
screen "Air System" 1280x800, template "Template"
   Button "Button_16" at 609,168 size 64x25; TextOn 'Alarm'; TextOff 'Text'
   Button "Button_2" at 602,168 size 71x25; TextOn 'Alarm'; TextOff 'Shutdown'
      Visibility <- "10 DI_DATA_E131_SHTDN"
   Button "HmiScreenItemData_1" at 1,1 size 150x43; TextOn 'Back'; TextOff 'Main Index'
      on Release: ActivateScreen("02 Main Index", 0)
   Button "Button_15" at 464,168 size 57x25; TextOn 'Enabled'; TextOff 'Disabled'
   TextField "Text field_14" at 307,171 size 158x18; Text 'I & A Air Compressor'
   TextField "Text field_15" at 464,146 size 60x18; Text 'Enabled'
   TextField "Text field_16" at 530,146 size 64x18; Text 'Running'
   TextField "Text field_18" at 601,145 size 78x18; Text 'Shutdown'
   Button "Button_1" at 530,168 size 57x25; TextOn 'Enabled'; TextOff 'Stopped'
   TextField "Text field_1" at 282,55 size 561x26; Text 'Instrument & Atomising Air Compressor Control (E-131)'
   TextField "Text field_32" at 464,168 size 57x25; Text 'Enabled'
      Visibility <- "14_DQ_Data_E131ControlOut"
   TextField "Text field_2" at 530,168 size 57x25; Text 'Running'
      Visibility <- "10 DI_DATA_E131_OK"
   GraphicIOField "Graphic I/O field_2" at 703,308 size 196x199; PictureList "IA Compressor_2"
      ProcessValue <- "82_To_HMI_CA Blower Animation"
   Gauge "Gauge_1" at 791,570 size 184x184; CaptionText 'Open'; UnitText '%'
      ProcessValue <- "12_AI_Data_CV403_SCALED"
   TextField "Text field_20" at 374,532 size 529x26; Text 'Combustion Air/Inert Gas Pressure Control (CV-403)'
   IOField "I/O field_16" at 516,441 size 74x25; FormatPattern 9999; Unit  RPM
      ProcessValue <- "12_AI_Data_E139_RPM_SCALED"
   IOField "I/O field_1" at 602,441 size 69x25; FormatPattern 999.99; Unit  A
      ProcessValue <- "12_AI_Data_E139_AMPS_SCALED"
   TextField "Text field_7" at 364,279 size 391x26; Text 'Combustion Air Blower Control (E-139)'
   Button "Button_3" at 464,395 size 57x25; TextOn 'Enabled'; TextOff 'Disabled'
   TextField "Text field_4" at 464,373 size 60x18; Text 'Enabled'
   TextField "Text field_5" at 624,373 size 40x18; Text 'Fault'
   Button "Button_5" at 615,396 size 57x25; TextOn 'Enabled'; TextOff 'Healthy'
   TextField "Text field_8" at 464,395 size 57x25; Text 'Enabled'
      Visibility <- "14_DQ_Data_E139_CNTRL"
   Button "Button_6" at 616,395 size 57x25; TextOn 'Alarm'; TextOff 'Fault'
      Visibility <- "10_DI_Data_E139_VSD_FLT"
      Appearance <- "10_DI_Data_E139_VSD_FLT"
   TextField "Text field_11" at 320,444 size 84x18; Text 'Motor RPM'
   TextField "Text field_3" at 307,399 size 124x18; Text 'Combustion Air'
   IOField "I/O field_5" at 429,441 size 75x25; Authorization "Operating Mode"; FormatPattern 9999; Unit  RPM
      ProcessValue <- "80_From_HMI_E139_SET_SPEED"
   Button "HmiScreenItemData_11" at 1016,173 size 69x51; TextOn 'RESET'; TextOff 'Reset'; Authorization "Operating Mode"
      on Press: function_b14e0dd5("82_To_HMI_I&A Compressor Reset Hours", 0)
   IOField "I/O field_8" at 941,175 size 65x25; FormatPattern 99999; Unit  h
      ProcessValue <- "82_To_HMI_I&A Compressor Run Hours(1)"
   IOField "I/O field_9" at 941,205 size 65x25; Authorization "Commissioning"; FormatPattern 99999; Unit  h
      ProcessValue <- "82_To_HMI_I&A Compressor Service Time Hours"
   TextField "Text field_19" at 911,174 size 37x20; Text 'Run'
   TextField "Text field_21" at 911,205 size 37x20; Text 'Set'
   TextField "Text field_13" at 954,78 size 140x20; Text 'Service Hour E131'
   Button "HmiScreenItemData_12" at 1016,428 size 69x51; TextOn 'RESET'; TextOff 'Reset'; Authorization "Operating Mode"
      on Press: function_b14e0dd5("82_To_HMI_CA Blower Reset Hours", 0)
   IOField "I/O field_10" at 941,427 size 65x25; FormatPattern 9999; Unit h
      ProcessValue <- "82_To_HMI_CA Blower Run Hours"
   IOField "I/O field_11" at 941,457 size 65x25; Authorization "Commissioning"; FormatPattern 9999; Unit  h
      ProcessValue <- "82_To_HMI_CA Blower Service Time Hours"
   TextField "Text field_22" at 911,429 size 37x20; Text 'Run'
   TextField "Text field_23" at 911,459 size 37x20; Text 'Set'
   TextField "Text field_24" at 954,329 size 148x20; Text 'Service Hours E139'
   Button "HmiScreenItemData_13" at 933,357 size 183x34; TextOn 'Back'; TextOff 'Text'
   IOField "I/O field_13" at 983,362 size 40x25; FormatPattern 99; Unit h
      ProcessValue <- "82_To_HMI_CA Blower Run Hours"
   IOField "I/O field_14" at 1025,362 size 40x25; FormatPattern 99; Unit m
      ProcessValue <- "82_To_HMI_CA Blower Run Minutes"
   IOField "I/O field_15" at 940,362 size 40x25; FormatPattern 99; Unit d
      ProcessValue <- "82_To_HMI_CA Blower Run Days"
   Button "HmiScreenItemData_14" at 928,105 size 183x34; TextOn 'Back'; TextOff 'Text'
   IOField "I/O field_17" at 978,109 size 40x25; FormatPattern 99; Unit h
      ProcessValue <- "82_To_HMI_I&A Compressor Run Hours"
   IOField "I/O field_18" at 1021,109 size 40x25; FormatPattern 99; Unit m
      ProcessValue <- "82_To_HMI_I&A Compressor Run Minutes"
   IOField "I/O field_19" at 1064,109 size 40x25; FormatPattern 99; Unit s
      ProcessValue <- "82_To_HMI_I&A Compressor Run Seconds"
   Button "Button_4" at 840,56 size 57x25; TextOn 'Alarm'; TextOff 'Service'
      Visibility <- "82_To_HMI_I&A Compressor Service Due"
   Button "Button_7" at 840,280 size 57x25; TextOn 'Alarm'; TextOff 'Service'
      Visibility <- "82_To_HMI_CA Blower Service Due"
   TextField "Text field_26" at 773,754 size 224x22; Text 'Modulating Valve Position'
   GraphicView "Graphic view_91" at 713,108 size 113x127; Picture "Graphic_246"
   GraphicIOField "Graphic I/O field_5" at 705,101 size 128x139; PictureList "New IA Compressor"
      ProcessValue <- "82_To_HMI_IA Compressor Animation"
      Visibility <- "68_Sys_Status_Data_IA_PRES_IN_RNG(1)"
   GraphicView "Graphic view_93" at 838,105 size 48x132; Picture "Graphic_248"
   GraphicView "Graphic view_2" at 823,160 size 19x12; Picture "Graphic_63"
   GraphicView "Graphic view_79" at 823,197 size 19x12; Picture "Graphic_63"
   Bar "Bar_1" at 852,115 size 20x105; Unit  %; MinimumValue 0; MaximumValue 100
      ProcessValue <- "12_AI_Data_PIT112In_SCALED"
      MaximumValue <- "84_Setpoints_PIT112_HighHigh"
   Button "HmiScreenItemData_4" at 1129,1 size 150x43; TextOn 'I&A Compressor Ok'; TextOff 'Back'
      on Release: function_efd93a16()
   IOField "I/O field_20" at 431,212 size 70x25; FormatPattern 99.99; Unit  Bar
      ProcessValue <- "12_AI_Data_PIT112In_SCALED"
   TextField "Text field_28" at 307,216 size 126x18; Text 'System Pressure'
   TextField "Text field_10" at 306,584 size 173x20; Text 'Air / Inert Gas Pressure'
   Button "Button_9" at 630,581 size 57x25; TextOn 'Enabled'; TextOff 'Text'
   TextField "Text field_17" at 306,620 size 310x20; Text 'Air / Inert Gas Pressure Setpoint (Pre-Ignition)'
   Button "Button_11" at 630,618 size 57x25; TextOn 'Enabled'; TextOff 'Text'
   TextField "Text field_12" at 311,736 size 182x20; Text 'Modulating Valve Position'
   TextField "Text field_25" at 306,657 size 310x20; Text 'Air / Inert Gas Pressure Setpoint (Post-Ignition)'
   Button "Button_10" at 630,655 size 57x25; TextOn 'Enabled'; TextOff 'Text'
   IOField "I/O field_2" at 625,582 size 66x25; FormatPattern 999; Unit  mbar
      ProcessValue <- "12_AI_Data_PIT402_SCALED"
   IOField "I/O field_3" at 625,618 size 66x25; Authorization "Commissioning"; FormatPattern 999; Unit  mbar
      ProcessValue <- "84_Setpoints_PIT402_Pilot_Target"
   IOField "I/O field_6" at 625,734 size 66x25; FormatPattern 999; Unit  %
      ProcessValue <- "16_AQ_Data_CV403_CNTRL"
   IOField "I/O field_7" at 625,692 size 66x23; FormatPattern 999; Unit  mBar
      ProcessValue <- "19_AUTO_CMNDS_Data_PIT402_Target"
      Appearance <- "19_AUTO_CMNDS_Data_PIT402_Target"
   IOField "I/O field_12" at 625,655 size 66x25; Authorization "Commissioning"; FormatPattern 999; Unit  mbar
      ProcessValue <- "84_Setpoints_PIT402_Main_Target"
   TextField "Text field_27" at 697,736 size 58x20; Text 'Opened'
   TextField "Text field_29" at 306,694 size 264x20; Text 'Air / Inert Gas Pressure Setpoint (Current)'
   AlarmView "Alarm view_1" at 0,777 size 1280x23
   TextField "Text field_6" at 531,373 size 64x18; Text 'Running'
   TextField "Text field_9" at 530,395 size 57x25; Text 'Running'
      Visibility <- "10_DI_Data_E139_RUNNING"
   IOField "I/O field_4" at 917,398 size 89x25; FormatPattern 999999; Unit h
      ProcessValue <- "82_To_HMI_CA Blower Total Run Hours"
   TextField "Text field_30" at 1011,400 size 123x20; Text 'Total Run Hours'
   IOField "I/O field_21" at 916,146 size 90x25; FormatPattern 999999; Unit  h
      ProcessValue <- "82_To_HMI_I&A Compressor Total Run Hours"
   TextField "Text field_31" at 1011,148 size 123x20; Text 'Total Run Hours'
   IOField "I/O field_22" at 935,109 size 40x25; FormatPattern 99; Unit d
      ProcessValue <- "82_To_HMI_P301 CSW Pump Run Days"
   IOField "I/O field_23" at 1068,362 size 40x25; FormatPattern 99; Unit s
      ProcessValue <- "82_To_HMI_CA Blower Run Seconds"

screen "Cooling System" 1280x800, template "Template"
   Group "Group_1" at 335,308 size 88x156; Picture "Graphic_148"
   Group "Group_2" at 298,412 size 194x121; Picture "Graphic_224"
   GraphicView "Graphic view_14" at 335,308 size 85x153; Picture "Graphic_148"
   GraphicView "Graphic view_9" at 298,414 size 189x119; Picture "Graphic_224"
   GraphicView "Graphic view_13" at 501,485 size 115x33; Picture "Graphic_232"
   GraphicView "Graphic view_1" at 446,429 size 75x87; Picture "Graphic_238"
   GraphicView "Graphic view_34" at 489,470 size 52x87; Picture "Graphic_169"
   GraphicView "Graphic view_11" at 80,468 size 424x50; Picture "Graphic_232"
   Group "Group_3" at 298,308 size 194x225; Picture "Graphic_148"
   GraphicView "Graphic view_2" at 480,389 size 43x49; Picture "Graphic_231"
   GraphicView "Graphic view_23" at 832,606 size 29x189; Picture "Graphic_231"
   GraphicView "Graphic view_18" at 802,567 size 88x52; Picture "Graphic_240"
   GraphicView "Graphic view_7" at 175,602 size 43x189; Picture "Graphic_231"
   GraphicView "Graphic view_29" at 964,565 size 56x50; Picture "Graphic_232"
   GraphicView "Graphic view_16" at 1150,564 size 56x50; Picture "Graphic_232"
   GraphicView "Graphic view_10" at 175,547 size 43x16; Picture "Graphic_231"
   GraphicView "Graphic view_8" at 25,514 size 207x209; Picture "Graphic_230"
   Button "HmiScreenItemData_1" at 1,1 size 150x43; TextOn 'Back'; TextOff 'Main Index'
      on Release: ActivateScreen("02 Main Index", 0)
   Rectangle "Rectangle_8" at 237,87 size 528x35
      Visibility <- "80_From_HMI_P301_PRSNT"
   Button "Button_15" at 468,92 size 57x25; TextOn 'Enabled'; TextOff 'Disabled'
      Visibility <- "80_From_HMI_P301_PRSNT"
   Button "Button_16" at 622,92 size 64x25; TextOn 'Alarm'; TextOff 'Text'
      Visibility <- "80_From_HMI_P301_PRSNT"
   TextField "Text field_14" at 239,94 size 185x20; Text 'Cooling Sea Water Pump'
   Button "Button_1" at 545,92 size 57x25; TextOn 'Enabled'; TextOff 'Stopped'
      Visibility <- "80_From_HMI_P301_PRSNT"
   Rectangle "Rectangle_1" at 236,83 size 530x212
      Visibility <- "80_From_HMI_P301_PRSNT"
   TextField "Text field_1" at 387,56 size 235x26; Text 'Cooling System Control'
   TextField "Text field_32" at 468,92 size 57x25; Text 'Enabled'
      Visibility <- "10 DI_DATA_P301_ENBLD"
   TextField "Text field_2" at 543,92 size 59x25; Text 'Running'
      Visibility <- "10_DI_Data_CV311_OPN(1)"
   Button "Button_2" at 622,92 size 64x25; TextOn 'Alarm'; TextOff 'Tripped'
      Visibility <- "10 DI_DATA_P301_TRIPPED"
      Appearance <- "10 DI_DATA_P301_TRIPPED"
   TextField "Text field_72" at 2,524 size 121x38; Text 'Cooling Seawater Inlet'
   GraphicView "Graphic view_17" at 464,297 size 75x99; Picture "Graphic_229"
   GraphicView "Graphic view_4" at 801,333 size 43x255; Picture "Graphic_231"
   GraphicView "Graphic view_5" at 786,305 size 72x46; Picture "Graphic_234"
   GraphicView "Graphic view_6" at 25,472 size 56x43; Picture "Graphic_235"
   TextField "Text field_7" at 12,598 size 58x20; Text 'CV-312'
   TextField "Text field_33" at 352,317 size 54x22; Text 'Closed'
      Visibility <- "10_DI_Data_CV311_CLSD"
   TextField "Text field_3" at 352,317 size 54x22; Text 'Opened'
      Visibility <- "10_DI_Data_CV311_OPN"
   TextField "Text field_71" at 351,343 size 58x20; Text 'CV-311'
   GraphicView "Graphic view_3" at 159,470 size 75x87; Picture "Graphic_239"
   TextField "Text field_5" at 534,295 size 105x38; Text 'To Inert Gas Generator'
   TextField "Text field_69" at 13,624 size 54x22; Text 'Closed'
      Visibility <- "10_DI_Data_CV312_CLSD"
   TextField "Text field_6" at 853,250 size 125x55; Text 'Warm Water From Inert Gas Generator'
   GraphicView "Graphic view_31" at 248,441 size 24x34; Picture "Graphic_36"
   TextField "Text field_17" at 230,422 size 62x20; Text 'PIT-359'
   IOField "I/O field_6" at 226,403 size 68x18; FormatPattern 99.99; Unit  Bar
      ProcessValue <- "12_AI_Data_PIT359_SCALED"
   GraphicView "Graphic view_21" at 849,377 size 88x52; Picture "Graphic_241"
   GraphicView "Graphic view_22" at 848,417 size 43x157; Picture "Graphic_231"
   TextField "Text field_8" at 867,659 size 78x55; Text 'Drain To Oily Bilge Tank'
   GraphicView "Graphic view_25" at 896,422 size 43x134; Picture "Graphic_231"
   GraphicView "Graphic view_26" at 898,526 size 73x87; Picture "Graphic_242"
   Group "Group_6" at 1006,404 size 194x225; Picture "Graphic_148"
   TextField "Text field_12" at 1053,439 size 58x20; Text 'CV-322'
   TextField "Text field_13" at 1054,413 size 54x22; Text 'Closed'
      Visibility <- "10_DI_Data_CV322_CLSD"
   TextField "Text field_19" at 1054,413 size 54x22; Text 'Opened'
      Visibility <- "10_DI_Data_CV322_OPN"
   TextField "Text field_20" at 1190,615 size 88x38; Text 'To Overboard'
   GraphicView "Graphic view_24" at 697,598 size 181x170; Picture "Graphic_230"
   TextField "Text field_9" at 681,704 size 58x20; Text 'CV-321'
   TextField "Text field_11" at 682,678 size 54x22; Text 'Closed'
      Visibility <- "10_DI_Data_CV321_CLSD"
   GraphicView "Graphic view_15" at 244,714 size 40x61; Picture "Graphic_236"
   TextField "Text field_21" at 214,658 size 93x55; Text 'To Existing Flue Gas Scrubber'
   TextField "Text field_70" at 13,624 size 54x22; Text 'Opened'
      Visibility <- "10_DI_Data_CV312_OPN"
   TextField "Text field_10" at 682,678 size 54x22; Text 'Opened'
      Visibility <- "10_DI_Data_CV321_OPN"
   GraphicView "Graphic view_32" at 512,546 size 30x121; Picture "Graphic_147"
   TextField "Text field_4" at 600,529 size 79x55; Text 'Cooling Seawater To GCU'
   GraphicView "Graphic view_19" at 624,477 size 56x43; Picture "Graphic_235"
   GraphicView "Graphic view_33" at 508,659 size 40x61; Picture "Graphic_236"
   TextField "Text field_22" at 481,722 size 79x55; Text 'Cooling Seawater To PGC'
   GraphicView "Graphic view_12" at 891,714 size 40x61; Picture "Graphic_236"
   GraphicView "Graphic view_30" at 1206,568 size 56x43; Picture "Graphic_235"
   GraphicView "Graphic view_35" at 803,244 size 40x61; Picture "Graphic_236"
   Button "HmiScreenItemData_4" at 1129,1 size 150x43; TextOn 'I&A Compressor Ok'; TextOff 'Back'
      on Release: function_efd93a16()
   AlarmView "Alarm view_1" at 0,777 size 1280x23
   Button "HmiScreenItemData_11" at 345,230 size 69x51; TextOn 'RESET'; TextOff 'Reset'; Authorization "Operating Mode"
      on Press: function_b14e0dd5("82_To_HMI_P301 CSW Pump Reset Hours", 0)
   IOField "I/O field_8" at 270,232 size 65x25; FormatPattern 99999; Unit  h
      ProcessValue <- "64_Functioning Hours_P301_IDB_Hours Functioning"
   IOField "I/O field_9" at 270,262 size 65x25; Authorization "Commissioning"; FormatPattern 99999; Unit  h
      ProcessValue <- "82_To_HMI_P301 CSW Pump Service Time Hours"
   TextField "Text field_23" at 240,231 size 37x20; Text 'Run'
   TextField "Text field_24" at 240,262 size 37x20; Text 'Set'
   TextField "Text field_25" at 283,121 size 141x20; Text 'Service Hour P301'
   Button "HmiScreenItemData_14" at 263,163 size 183x34; TextOn 'Back'; TextOff 'Text'
   IOField "I/O field_17" at 312,167 size 40x25; FormatPattern 99; Unit h
      ProcessValue <- "82_To_HMI_P301 CSW Pump Run Hours"
   IOField "I/O field_18" at 355,167 size 40x25; FormatPattern 99; Unit m
      ProcessValue <- "82_To_HMI_P301 CSW Pump Run Minutes"
   IOField "I/O field_19" at 398,167 size 40x25; FormatPattern 99; Unit s
      ProcessValue <- "82_To_HMI_P301 CSW Pump Run Seconds"
   IOField "I/O field_21" at 245,203 size 90x25; FormatPattern 999999; Unit  h
      ProcessValue <- "82_To_HMI_P301 CSW Pump Total Run Hours"
   TextField "Text field_31" at 340,205 size 123x20; Text 'Total Run Hours'
   Button "Button_17" at 701,92 size 57x25; TextOn 'Alarm'; TextOff 'Service'
      Visibility <- "80_From_HMI_P301_PRSNT"
   Button "Button_9" at 701,92 size 57x25; TextOn 'Alarm'; TextOff 'Service'
      Visibility <- "82_To_HMI_P301 CSW Pump Service Due"
   IOField "I/O field_1" at 270,167 size 40x25; FormatPattern 99; Unit d
      ProcessValue <- "82_To_HMI_P301 CSW Pump Run Days"
   Rectangle "Rectangle_7" at 224,48 size 554x250
      Visibility <- "80_From_HMI_P301_PRSNT"
   Button "HmiScreenItemData_2" at 520,167 size 184x67; TextOn 'FRESH WATER SYSTEM'; TextOff 'Fresh Water System'; Authorization "Operating Mode"
      on Release: ActivateScreen("Fresh Water System", 0)
      Visibility <- "80_From_HMI_P305_PRSNT"
   Button "HmiScreenItemData_3" at 595,392 size 170x41; TextOn 'STOP CSW OVERRUN'; TextOff 'Stop CSW Overrun'; Authorization "Operating Mode"
      on Press: function_b14e0dd5("80_From_HMI_CSW OVR Stop", 0)
      Appearance <- "10_DI_Data_CV311_OPN"
   Group "Group_4" at 1043,404 size 88x156; Picture "Graphic_148"
   Group "Group_5" at 1006,508 size 194x121; Picture "Graphic_224"
   GraphicView "Graphic view_27" at 1043,404 size 85x153; Picture "Graphic_148"
   GraphicView "Graphic view_28" at 1006,511 size 189x119; Picture "Graphic_224"

screen "Fuel System" 1280x800, template "Template"
   GraphicView "Graphic view_4" at 570,430 size 24x23; Picture "Graphic_102"
   Button "HmiScreenItemData_1" at 1,1 size 150x43; TextOn 'Back'; TextOff 'Main Index'
      on Release: ActivateScreen("02 Main Index", 0)
   TextField "Text field_3" at 691,522 size 55x18; Text 'E-500B'
   GraphicView "Graphic view_16" at 658,375 size 123x15; Picture "Graphic_99"
   GraphicIOField "Graphic I/O field_1" at 686,356 size 60x65; PictureList "Pump Ani"
      ProcessValue <- "82_To_HMI_Fuel Pump 1 Animation"
   GraphicView "Graphic view_10" at 657,477 size 124x15; Picture "Graphic_99"
   GraphicIOField "Graphic I/O field_2" at 686,459 size 60x65; PictureList "Pump Ani"
      ProcessValue <- "82_To_HMI_Fuel Pump 2 Animation"
   GraphicView "Graphic view_17" at 642,390 size 15x94; Picture "Graphic_101"
   GraphicView "Graphic view_14" at 643,466 size 21x25; Picture "Graphic_96"
   GraphicView "Graphic view_18" at 643,376 size 24x23; Picture "Graphic_102"
   GraphicView "Graphic view_19" at 638,425 size 18x23; Picture "Graphic_105"
   GraphicView "Graphic view_20" at 782,390 size 15x94; Picture "Graphic_101"
   GraphicView "Graphic view_9" at 772,376 size 24x23; Picture "Graphic_104"
   GraphicView "Graphic view_21" at 771,467 size 25x24; Picture "Graphic_97"
   GraphicView "Graphic view_7" at 783,426 size 19x24; Picture "Graphic_103"
   GraphicView "Graphic view_22" at 578,429 size 71x15; Picture "Graphic_99"
   GraphicView "Graphic view_23" at 789,430 size 94x15; Picture "Graphic_99"
   GraphicView "Graphic view_24" at 672,375 size 18x15; Picture "Graphic_99"
   GraphicView "Graphic view_25" at 672,477 size 18x15; Picture "Graphic_99"
   TextField "Text field_2" at 691,422 size 56x18; Text 'E-500A'
   GraphicView "Graphic view_1" at 621,429 size 27x15; Picture "Graphic_99"
   Button "Button_15" at 157,172 size 57x25; TextOn 'Enabled'; TextOff 'Disabled'
   TextField "Text field_14" at 59,174 size 92x20; Text 'Fuel Pump 1'
   TextField "Text field_15" at 161,151 size 60x18; Text 'Enabled'
   TextField "Text field_18" at 391,149 size 87x18; Text 'Service Due'
   Button "Button_17" at 396,172 size 57x25; TextOn 'Alarm'; TextOff 'Service'
   Button "Button_18" at 159,375 size 57x25; TextOn 'Enabled'; TextOff 'Disabled'
   TextField "Text field_19" at 61,377 size 92x20; Text 'Fuel Pump 2'
   Button "Button_20" at 398,375 size 57x25; TextOn 'Alarm'; TextOff 'Service'
   Rectangle "Rectangle_13" at 678,350 size 77x92
      Appearance <- "10_DI_Data_E500A_TRIPPED"
   Rectangle "Rectangle_14" at 678,453 size 77x92
      Appearance <- "10_DI_Data_E500B_TRIPPED(1)"
   TextField "Text field_7" at 678,544 size 83x18; Text 'Duty Pump'
      Visibility <- "101_Fuel_Pumps_DB_Duty Is B"
   TextField "Text field_12" at 678,333 size 83x18; Text 'Duty Pump'
      Visibility <- "101_Fuel_Pumps_DB_Duty Is A"
   GraphicView "Graphic view_8" at 854,430 size 152x15; Picture "Graphic_99"
   Button "Button_9" at 396,172 size 57x25; TextOn 'Alarm'; TextOff 'Service'
      Visibility <- "82_To_HMI_E500A Fuel Pump Service Due"
   Button "Button_10" at 398,375 size 57x25; TextOn 'Alarm'; TextOff 'Service'
      Visibility <- "82_To_HMI_E500B Fuel Pump Service Due"
   GraphicView "Graphic view_76" at 951,407 size 20x26; Picture "Graphic_36"
   TextField "Text field_23" at 933,442 size 61x18; Text 'PIT-204'
   GraphicView "Graphic view_46" at 997,420 size 20x24; Picture "Graphic_40"
   GraphicView "Graphic view_54" at 1016,372 size 24x21; Picture "Graphic_107"
   TextField "Text field_33" at 1022,392 size 60x18; Text 'TIT-202'
   GraphicView "Graphic view_45" at 1005,315 size 13x117; Picture "Graphic_57"
   TextField "Text field_1" at 1049,301 size 172x18; Text 'IGG Pilot & Main Burner'
   GraphicView "Graphic view_2" at 1006,305 size 20x23; Picture "Graphic_102"
   GraphicView "Graphic view_3" at 549,738 size 6x20; Picture "Graphic_113"
   GraphicView "Graphic view_5" at 557,731 size 25x24; Picture "Graphic_111"
   GraphicView "Graphic view_66" at 568,552 size 15x192; Picture "Graphic_112"
   GraphicView "Graphic view_6" at 568,442 size 15x192; Picture "Graphic_112"
   GraphicView "Graphic view_11" at 551,740 size 15x15; Picture "Graphic_99"
   Button "Button_13" at 157,172 size 57x25; TextOn 'Enabled'; TextOff 'Enabled'
      Visibility <- "10_DI_Data_E500A_ENBLD(1)"
   Button "Button_14" at 159,375 size 57x25; TextOn 'Enabled'; TextOff 'Enabled'
      Visibility <- "10_DI_Data_E500B_ENBLD(1)"
   Button "HmiScreenItemData_7" at 525,369 size 69x51; TextOn 'Back'; TextOff 'PSelect'; Authorization "Operating Mode"
      on Press: function_b14e0dd5("80_From_HMI_SW_DTY_PMP_E500", 0)
   IOField "I/O field_1" at 934,390 size 65x22; FormatPattern 99.99; Unit  Bar
      ProcessValue <- "12_AI_Data_PIT204In_SCALED"
   IOField "I/O field_3" at 312,171 size 65x25; FormatPattern 999999
      ProcessValue <- "64_Functioning Hours_E500A_IDB_Hours Functioning"
   TextField "Text field_5" at 315,149 size 72x18; Text 'Hour Run'
   IOField "I/O field_6" at 314,374 size 65x25; FormatPattern 999999
      ProcessValue <- "64_Functioning Hours_E500B_IDB_Hours Functioning"
   Button "Button_1" at 233,172 size 57x25; TextOn 'Alarm'; TextOff 'Text'
   TextField "Text field_6" at 241,149 size 45x18; Text 'Alarm'
   Button "Button_2" at 235,375 size 57x25; TextOn 'Alarm'; TextOff 'Text'
   Button "Button_3" at 233,172 size 57x25; TextOn 'Alarm'; TextOff 'Tripped'
      Visibility <- "10_DI_Data_E500A_TRIPPED"
      Appearance <- "10_DI_Data_E500A_TRIPPED"
   Button "Button_4" at 235,375 size 57x25; TextOn 'Alarm'; TextOff 'Tripped'
      Visibility <- "10_DI_Data_E500B_TRIPPED(1)"
      Appearance <- "10_DI_Data_E500B_TRIPPED(1)"
   IOField "I/O field_4" at 1043,373 size 55x18; FormatPattern 99.9; Unit  °C
      ProcessValue <- "12_AI_Data_TIT202In_SCALED"
   Button "HmiScreenItemData_3" at 1129,1 size 150x43; TextOn 'I&A Compressor Ok'; TextOff 'Back'
      on Release: function_efd93a16()
   AlarmView "Alarm view_1" at 0,777 size 1280x23
   Button "HmiScreenItemData_11" at 253,294 size 69x51; TextOn 'RESET'; TextOff 'Reset'; Authorization "Operating Mode"
      on Press: function_b14e0dd5("82_To_HMI_E500A Fuel Pump Reset Hours", 0)
   IOField "I/O field_8" at 178,296 size 65x25; FormatPattern 99999; Unit  h
      ProcessValue <- "64_Functioning Hours_E500A_IDB_Hours Functioning"
   IOField "I/O field_9" at 178,326 size 65x25; Authorization "Commissioning"; FormatPattern 99999; Unit  h
      ProcessValue <- "82_To_HMI_E500A Fuel Pump Service Time Hours"
   TextField "Text field_8" at 148,295 size 37x20; Text 'Run'
   TextField "Text field_21" at 148,326 size 37x20; Text 'Set'
   TextField "Text field_13" at 191,201 size 151x20; Text 'Service Hour E500A'
   Button "HmiScreenItemData_14" at 171,227 size 150x34; TextOn 'Back'; TextOff 'Text'
   IOField "I/O field_17" at 176,231 size 54x25; FormatPattern 999; Unit h
      ProcessValue <- "64_Functioning Hours_E500A_IDB_Hours Functioning"
   IOField "I/O field_18" at 232,231 size 40x25; FormatPattern 99; Unit m
      ProcessValue <- "82_To_HMI_E500A Fuel Pump Run Minutes"
   IOField "I/O field_19" at 275,231 size 40x25; FormatPattern 99; Unit s
      ProcessValue <- "82_To_HMI_E500A Fuel Pump Run Seconds"
   IOField "I/O field_21" at 153,267 size 90x25; FormatPattern 999999; Unit  h
      ProcessValue <- "82_To_HMI_E500A Fuel Pump Total Run Hours"
   TextField "Text field_31" at 248,269 size 123x20; Text 'Total Run Hours'
   Button "HmiScreenItemData_2" at 255,502 size 69x51; TextOn 'RESET'; TextOff 'Reset'; Authorization "Operating Mode"
      on Press: function_b14e0dd5("82_To_HMI_E500B Fuel Pump Reset Hours", 0)
   IOField "I/O field_5" at 180,504 size 65x25; FormatPattern 99999; Unit  h
      ProcessValue <- "64_Functioning Hours_E500B_IDB_Hours Functioning"
   IOField "I/O field_7" at 180,534 size 65x25; Authorization "Commissioning"; FormatPattern 99999; Unit  h
      ProcessValue <- "82_To_HMI_E500B Fuel Pump Service Time Hours"
   TextField "Text field_9" at 150,503 size 37x20; Text 'Run'
   TextField "Text field_10" at 150,534 size 37x20; Text 'Set'
   TextField "Text field_11" at 193,402 size 149x20; Text 'Service Hour E500B'
   Button "HmiScreenItemData_4" at 174,430 size 150x34; TextOn 'Back'; TextOff 'Text'
   IOField "I/O field_10" at 179,434 size 54x25; FormatPattern 999; Unit h
      ProcessValue <- "64_Functioning Hours_E500B_IDB_Hours Functioning"
   IOField "I/O field_11" at 235,434 size 40x25; FormatPattern 99; Unit m
      ProcessValue <- "82_To_HMI_E500B Fuel Pump Run Minutes"
   IOField "I/O field_12" at 278,434 size 40x25; FormatPattern 99; Unit s
      ProcessValue <- "82_To_HMI_E500B Fuel Pump Run Seconds"
   IOField "I/O field_13" at 155,475 size 90x25; FormatPattern 999999; Unit  h
      ProcessValue <- "82_To_HMI_E500B Fuel Pump Total Run Hours"
   TextField "Text field_16" at 250,477 size 123x20; Text 'Total Run Hours'

screen "IG Transfer Mode" 1280x800, template "Template"
   Group "Group_1" at 596,282 size 37x72; Picture "Graphic_148"
   Group "Group_2" at 581,330 size 80x56; Picture "Graphic_224"
   GraphicView "Graphic view_14" at 596,282 size 36x71; Picture "Graphic_148"
   GraphicView "Graphic view_9" at 581,331 size 78x55; Picture "Graphic_224"
   Group "Group_4" at 670,65 size 37x72; Picture "Graphic_148"
   Group "Group_5" at 655,113 size 80x56; Picture "Graphic_224"
   GraphicView "Graphic view_28" at 670,65 size 36x71; Picture "Graphic_148"
   GraphicView "Graphic view_29" at 655,114 size 78x55; Picture "Graphic_224"
   Group "Group_7" at 302,283 size 37x72; Picture "Graphic_148"
   Group "Group_8" at 287,331 size 80x56; Picture "Graphic_224"
   GraphicView "Graphic view_7" at 302,283 size 36x71; Picture "Graphic_148"
   GraphicView "Graphic view_10" at 287,332 size 78x55; Picture "Graphic_224"
   GraphicView "Graphic view_6" at 871,216 size 36x71; Picture "Graphic_148"
   Group "Group_10" at 871,216 size 37x72; Picture "Graphic_148"
   Group "Group_11" at 856,264 size 80x56; Picture "Graphic_224"
   GraphicView "Graphic view_12" at 856,265 size 78x55; Picture "Graphic_224"
   GraphicView "Graphic view_24" at 761,309 size 18x78; Picture "Graphic_231"
   GraphicView "Graphic view_27" at 472,141 size 336x19; Picture "Graphic_232"
   Group "Group_6" at 655,65 size 80x104; Picture "Graphic_148"
   GraphicView "Graphic view_8" at 454,142 size 31x33; Picture "Graphic_178"
   Group "Group_3" at 581,282 size 80x104; Picture "Graphic_148"
   Button "HmiScreenItemData_1" at 1,1 size 150x43; TextOn 'Back'; TextOff 'Main Index'
      on Release: ActivateScreen("02 Main Index", 0)
   TextField "Text field_5" at 111,336 size 84x55; Text 'From Inert Gas Generator'
   TextField "Text field_12" at 655,72 size 58x20; Text 'CV-432'
   TextField "Text field_13" at 656,48 size 54x22; Text 'Closed'
      Visibility <- "10_DI_Data_CV432_CLSD"
   TextField "Text field_19" at 656,48 size 54x22; Text 'Opened'
      Visibility <- "10_DI_Data_CV432_OPN"
   TextField "Text field_9" at 582,291 size 58x20; Text 'CV-431'
   TextField "Text field_10" at 583,268 size 54x22; Text 'Opened'
      Visibility <- "10_DI_Data_CV431_OPN"
   Button "HmiScreenItemData_17" at 1,46 size 150x43; TextOn 'IGG Plant'; TextOff 'IGGS Plant'
      on Release: ActivateScreen("Inert Gas Generator Plant", 0)
   GraphicView "Graphic view_35" at 696,328 size 264x286; Picture "Graphic_251"
   GraphicView "Graphic view_4" at 749,359 size 30x28; Picture "Graphic_169"
   GraphicView "Graphic view_18" at 759,509 size 25x27; Picture "Graphic_265"
   GraphicView "Graphic view_20" at 759,531 size 35x38; Picture "Graphic_266"
   GraphicView "Graphic view_5" at 992,464 size 168x269; Picture "Graphic_150"
   GraphicView "Graphic view_21" at 773,548 size 216x22; Picture "Graphic_232"
   GraphicView "Graphic view_22" at 976,533 size 20x49; Picture "Graphic_271"
   GraphicView "Graphic view_23" at 1165,476 size 35x22; Picture "Graphic_232"
   GraphicView "Graphic view_25" at 1154,465 size 20x43; Picture "Graphic_271"
   GraphicView "Graphic view_26" at 640,358 size 115x17; Picture "Graphic_232"
   GraphicView "Graphic view_1" at 265,360 size 329x17; Picture "Graphic_232"
   GraphicView "Graphic view_17" at 453,166 size 18x202; Picture "Graphic_231"
   GraphicView "Graphic view_3" at 214,351 size 56x35; Picture "Graphic_279"
   Group "Group_9" at 287,283 size 80x104; Picture "Graphic_148"
   TextField "Text field_49" at 294,291 size 56x18; Text 'CV-401'
   TextField "Text field_50" at 292,268 size 54x22; Text 'Closed'
      Visibility <- "10_DI_Data_CV401_CLSD"
   TextField "Text field_51" at 292,268 size 54x22; Text 'Opened'
      Visibility <- "10_DI_Data_CV401_OPN"
   GraphicView "Graphic view_2" at 791,129 size 20x43; Picture "Graphic_280"
   TextField "Text field_1" at 874,131 size 88x38; Text 'To Cargo Blanketing'
   GraphicView "Graphic view_11" at 816,134 size 56x35; Picture "Graphic_279"
   TextField "Text field_48" at 744,627 size 112x20; Text 'PG Compressor'
      Appearance <- "10_DI_DATA_E_400_NOK"
   TextField "Text field_56" at 1202,508 size 71x18; Text 'For BWTS'
   TextField "Text field_2" at 1068,752 size 38x20; Text 'GCU'
   TextField "Text field_11" at 583,268 size 54x22; Text 'Closed'
      Visibility <- "10_DI_Data_CV431_CLSD"
   Button "HmiScreenItemData_3" at 1129,1 size 150x43; TextOn 'I&A Compressor Ok'; TextOff 'Back'
      on Release: function_efd93a16()
   AlarmView "Alarm view_1" at 0,777 size 1280x23
   GraphicView "Graphic view_83" at 1184,463 size 96x48; Picture "Graphic_235"
   Button "HmiScreenItemData_5" at 1165,453 size 114x70; TextOn 'Back'; TextOff 'Text'
      on Press: ActivateScreen("Balast Water Treatment Plant", 0)
   GraphicView "Graphic view_108" at 6,137 size 95x48; Picture "Left Arow"
   Button "HmiScreenItemData_14" at 5,124 size 106x107; TextOn 'Back'; TextOff 'Text'
      on Press: ActivateScreen("Inert Gas Generator Plant", 0)
   TextField "Text field_21" at 12,193 size 77x34; Text 'Inert Gas Generator'
   GraphicView "Graphic view_13" at 773,292 size 245x19; Picture "Graphic_232"
   GraphicView "Graphic view_15" at 762,293 size 31x33; Picture "Graphic_178"
   GraphicView "Graphic view_16" at 996,280 size 20x43; Picture "Graphic_280"
   TextField "Text field_3" at 1077,283 size 71x38; Text 'Ambient Air Inlet'
   GraphicView "Graphic view_19" at 1021,285 size 56x35; Picture "left small arrow"
   Group "Group_12" at 856,216 size 80x104; Picture "Graphic_148"
   Button "Button_1" at 666,321 size 296x306; TextOff 'Text'
      on Press: ActivateScreen("Inert Gas Conditioning Plant", 0)
   TextField "Text field_4" at 862,225 size 56x18; Text 'CV-441'
   TextField "Text field_6" at 862,202 size 54x22; Text 'Closed'
      Visibility <- "10_DI_DATA_CV441_CLSD"
   TextField "Text field_7" at 862,202 size 54x22; Text 'Opened'
      Visibility <- "10_DI_DATA_CV441_OPN"

screen "O2 Content Monitoring" 1280x800, template "Template"
   TextField "Text field_10" at 20,573 size 128x20; Text 'E600 O2 Content'
   Button "Button_9" at 180,571 size 57x25; TextOn 'Enabled'; TextOff 'Text'
   TextField "Text field_17" at 20,601 size 125x52; Text 'BWT O2 Content Setpoint'
   Button "Button_11" at 180,607 size 57x25; TextOn 'Enabled'; TextOff 'Text'
   TextField "Text field_20" at 153,468 size 171x26; Text 'E600 O2 Content'
   TextField "Text field_12" at 19,646 size 154x20; Text 'Cargo Blanketing O2'
   IOField "I/O field_2" at 177,571 size 74x25; FormatPattern s99.999; Unit %
      ProcessValue <- "12_AI_Data_E600O2ContentIn"
   IOField "I/O field_6" at 180,645 size 66x25; Authorization "Parameter Change"; FormatPattern 99.99; Unit  %
      ProcessValue <- "84_Setpoints_E600_CB_Target"
   TextField "Text field_3" at 484,512 size 160x20; Text 'Burner Fuel Pressure'
   Button "Button_3" at 644,510 size 57x25; TextOn 'Enabled'; TextOff 'Text'
   TextField "Text field_4" at 484,541 size 161x52; Text 'Burner Fuel Pressure Setpoint'
   TextField "Text field_5" at 575,468 size 296x26; Text 'Burner Fuel Control (CV-203)'
   TextField "Text field_6" at 483,585 size 110x20; Text 'Valve Position'
   IOField "I/O field_1" at 642,510 size 71x25; FormatPattern 99.99; Unit  bar
      ProcessValue <- "12_AI_Data_PIT205In_SCALED"
   IOField "I/O field_5" at 642,584 size 71x25; FormatPattern 999.99; Unit  %
      ProcessValue <- "16_AQ_Data_CV203_CNTRL"
   IOField "I/O field_3" at 180,607 size 66x25; Authorization "Parameter Change"; FormatPattern 99.99; Unit %
      ProcessValue <- "84_Setpoints_E600_BWT_Target"
   Button "HmiScreenItemData_3" at 1,1 size 150x43; TextOn 'Back'; TextOff 'Main Index'
      on Release: ActivateScreen("02 Main Index", 0)
   Button "HmiScreenItemData_1" at 1129,1 size 150x43; TextOn 'I&A Compressor Ok'; TextOff 'Back'
      on Release: function_efd93a16()
   AlarmView "Alarm view_1" at 0,777 size 1280x23
   Gauge "Gauge_2" at 258,545 size 210x210; UnitText '%'; CaptionText 'O2 Content'
      Visibility <- "80_From_HMI_CRG_BLNK_MODE"
      ProcessValue <- "12_AI_Data_E600O2ContentIn"
      MaximumValue <- "84_Setpoints_E600_CB_HighHigh"
   TextField "Text field_11" at 975,675 size 257x27; Text 'Proportionate Component PID'
   TextField "Text field_15" at 975,709 size 257x27; Text 'Integrative Component PID'
   TextField "Text field_16" at 975,742 size 257x27; Text 'Derivative Component PID'
   TextField "Text field_19" at 975,553 size 153x27; Text 'Derivation Time'
   TextField "Text field_1" at 977,490 size 153x27; Text 'GAIN'
   TextField "Text field_18" at 975,519 size 153x27; Text 'Integration Time'
   TextField "Text field_2" at 977,588 size 153x27; Text 'Maximum opening'
   Group "Group_16" at 1130,554 size 112x34; Authorization "User administration"; Picture "Graphic_284"; FormatPattern 99
   Switch "Switch_8" at 1223,676 size 32x29; CaptionText 'Switch'; TextOn 'ON'; TextOff 'OFF'; Authorization "User administration"; PictureOff "Design_5_PilotLight_Green_Off"; PictureOn "Design_5_PilotLight_Green_On"
      on Change: InvertBit("84_Setpoints_P_ON")
      ProcessValue <- "84_Setpoints_P_ON"
   Group "Group_15" at 1130,519 size 112x34; Authorization "User administration"; Picture "Graphic_284"; FormatPattern 99
   Switch "Switch_9" at 1223,710 size 32x29; CaptionText 'Switch'; TextOn 'ON'; TextOff 'OFF'; Authorization "User administration"; PictureOff "Design_5_PilotLight_Green_Off"; PictureOn "Design_5_PilotLight_Green_On"
      on Change: InvertBit("84_Setpoints_I_ON")
      ProcessValue <- "84_Setpoints_I_ON"
   Group "Group_3" at 1130,484 size 112x34; Authorization "User administration"; Picture "Graphic_284"; FormatPattern 99
   Switch "Switch_10" at 1223,741 size 32x29; CaptionText 'Switch'; TextOn 'ON'; TextOff 'OFF'; Authorization "User administration"; PictureOff "Design_5_PilotLight_Green_Off"; PictureOn "Design_5_PilotLight_Green_On"
      on Change: InvertBit("84_Setpoints_D_ON")
      ProcessValue <- "84_Setpoints_D_ON"
   Group "Group_1" at 1130,622 size 112x34; Authorization "User administration"; Picture "Graphic_284"; FormatPattern 99
   TextField "Text field_21" at 977,622 size 153x27; Text 'Minimum opening'
   Circle "Circle_29" at 30,726 size 20x20
      Appearance <- "Evolving Setpoint_DB_LevelBetter"
   TextField "Text field_22" at 59,722 size 217x27; Text 'O2 content closing Setpoint'
   TrendView "Trend view_1" at 13,53 size 1256x405
      Visibility <- "80_From_HMI_CRG_BLNK_MODE"
      ValueAxis2End <- "84_Setpoints_Max Opening"
      ValueAxis2Begin <- "84_Setpoints_Min Opening"
      ValueAxis1End <- "84_Setpoints_E600_CB_HighHigh"
   TrendView "Trend view_2" at 14,53 size 1259x409
      Visibility <- "80_From_HMI_BWT_BYPASS"
      ValueAxis2End <- "84_Setpoints_Max Opening"
      ValueAxis2Begin <- "84_Setpoints_Min Opening"
      ValueAxis1End <- "84_Setpoints_E600_BWT_HighHigh"
   Gauge "Gauge_3" at 258,545 size 210x210; UnitText '%'; CaptionText 'O2 Content'
      Visibility <- "80_From_HMI_BWT_BYPASS"
      ProcessValue <- "12_AI_Data_E600O2ContentIn"
      MaximumValue <- "84_Setpoints_E600_BWT_HighHigh"
   TextField "Text field_7" at 485,632 size 176x20; Text 'Atomising Air Pressure'
   Button "Button_1" at 650,630 size 57x25; TextOn 'Enabled'; TextOff 'Text'
   TextField "Text field_8" at 485,667 size 180x36; Text 'Pilot Air Press Setpoint'
   Button "Button_2" at 649,666 size 57x25; TextOn 'Enabled'; TextOff 'Text'
   TextField "Text field_9" at 484,742 size 110x20; Text 'Valve Position'
   IOField "I/O field_4" at 642,630 size 71x25; FormatPattern 99.99; Unit  bar
      ProcessValue <- "12_AI_Data_PIT113In_SCALED"
   IOField "I/O field_7" at 642,741 size 71x25; FormatPattern 999.99; Unit  %
      ProcessValue <- "16_AQ_Data_CV111_CNTRL"
   IOField "I/O field_8" at 642,666 size 71x25; Authorization "Commissioning"; FormatPattern 99.99; Unit  bar
      ProcessValue <- "84_Setpoints_PIT113_Pilot_Target"
   Group "Group_2" at 1130,588 size 112x34; Authorization "User administration"; Picture "Graphic_284"; FormatPattern 99
   IOField "I/O field_9" at 642,547 size 71x25; Authorization "Commissioning"; FormatPattern 99.99; Unit  bar
      ProcessValue <- "84_Setpoints_PIT205_Target"
   TextField "Text field_13" at 485,704 size 197x36; Text 'Burner Air Press Setpoint'
   Button "Button_4" at 649,703 size 57x25; TextOn 'Enabled'; TextOff 'Text'
   IOField "I/O field_10" at 642,703 size 71x25; Authorization "Commissioning"; FormatPattern 99.99; Unit  bar
      ProcessValue <- "84_Setpoints_PIT113_Burner_Target"
   Gauge "Gauge_4" at 721,547 size 211x211; UnitText '%'; CaptionText 'CV 203'
      ProcessValue <- "16_AQ_Data_CV203_CNTRL"
   GraphicView "Graphic view_22" at 1130,519 size 112x34; Picture "Graphic_284"
   IOField "D5_I/O field_2" at 1145,527 size 62x18; Authorization "User administration"; FormatPattern 99999
      ProcessValue <- "84_Setpoints_Integration Time"
   TextField "D5_Text field_2" at 1205,527 size 23x18; Text 'ms / km/h'
   GraphicView "Graphic view_23" at 1130,554 size 112x34; Picture "Graphic_284"
   IOField "D5_I/O field_3" at 1145,562 size 62x18; Authorization "User administration"; FormatPattern 99999
      ProcessValue <- "84_Setpoints_Derive Time"
   TextField "D5_Text field_3" at 1205,562 size 23x18; Text 'ms / km/h'
   GraphicView "Graphic view_25" at 1130,484 size 112x34; Picture "Graphic_284"
   IOField "D5_I/O field_10" at 1145,492 size 62x18; Authorization "User administration"; FormatPattern 99.9999
      ProcessValue <- "84_Setpoints_Gain"
   TextField "D5_Text field_10" at 1205,492 size 23x18; Text 'km/h'
   GraphicView "Graphic view_1" at 1130,622 size 112x34; Picture "Graphic_284"
   IOField "D5_I/O field_1" at 1145,630 size 62x18; Authorization "User administration"; FormatPattern 999; Unit %
      ProcessValue <- "84_Setpoints_Min Opening"
   TextField "D5_Text field_1" at 1205,630 size 23x18; Text 'km/h'
   GraphicView "Graphic view_2" at 1130,588 size 112x34; Picture "Graphic_284"
   IOField "D5_I/O field_5" at 1145,596 size 62x18; Authorization "User administration"; FormatPattern 999; Unit %
      ProcessValue <- "84_Setpoints_Max Opening"
   TextField "D5_Text field_5" at 1205,596 size 23x18; Text 'km/h'

PopupScreen "CV 203 Grafics" 810x675
   Button "Button_1" at 753,0 size 56x38; TextOff 'Text'; PictureOff "Graphic_286"
      on Click: function_efd93a16("CV 203 Grafics", 0, 0, -1, -1, 1)
   GraphicView "Graphic view_2" at 2,2 size 751x35; Picture "Graphic_287"
   TextField "Text field_1" at 285,7 size 229x26; Text 'O2 FUEL MODULATION'
   TrendView "Trend view_2" at 1,38 size 808x636
      Visibility <- "80_From_HMI_CRG_BLNK_MODE"
      ValueAxis2End <- "84_Setpoints_Max Opening"
      ValueAxis2Begin <- "84_Setpoints_Min Opening"
      ValueAxis1End <- "84_Setpoints_E600_CB_HighHigh"
   TrendView "Trend view_1" at 2,40 size 804x635
      Visibility <- "80_From_HMI_BWT_BYPASS"
      ValueAxis2End <- "84_Setpoints_Max Opening"
      ValueAxis2Begin <- "84_Setpoints_Min Opening"
      ValueAxis1End <- "84_Setpoints_E600_BWT_HighHigh"

PopupScreen "CV 403 Grafics" 810x675
   Button "Button_1" at 753,0 size 56x40; TextOff 'Text'; PictureOff "Graphic_286"
      on Click: function_efd93a16("CV 403 Grafics", 0, 0, -1, -1, 1)
   GraphicView "Graphic view_2" at 2,2 size 751x35; Picture "Graphic_287"
   TextField "Text field_1" at 285,9 size 281x26; Text 'IG PRESSURE MODULATION'
   TrendView "Trend view_2" at 1,39 size 809x635

screen "Commissioning Main Page" 1280x800, template "Template"
   on GenerateScreen: "TitleUpdater"()
   Button "HmiScreenItemData_1" at 1,2 size 150x43; TextOn 'Back'; TextOff 'Main Index'
      on Release: ActivateScreen("02 Main Index", 0)
   AlarmView "Alarm view_1" at 0,777 size 1280x23
   Button "HmiScreenItemData_4" at 790,100 size 200x35; TextOn 'Back'; TextOff 'BWT Settings'
   Button "Button_22" at 800,150 size 180x50; TextOff 'Target Setpoints'; Authorization "Commissioning"
      on Press: ActivateScreen("BWT Target Setpoints", 0)
   Button "Button_24" at 800,220 size 180x50; TextOff 'Process Times'; Authorization "Commissioning"
      on Press: ActivateScreen("BWT Process Times", 0)
   Button "HmiScreenItemData_3" at 540,100 size 200x35; TextOn 'Back'; TextOff 'GCU Settings'
   Button "Button_13" at 550,150 size 180x50; TextOff 'Digital Inputs'; Authorization "Commissioning"
      on Click: ActivateScreen("GCU Digital Inputs", 0)
   Button "Button_14" at 550,220 size 180x50; TextOff 'Digital Outputs'; Authorization "Operating Mode"
      on Click: ActivateScreen("GCU Digital Outputs", 0)
   Button "Button_15" at 550,290 size 180x50; TextOff 'Analogue Inputs'; Authorization "Commissioning"
      on Press: ActivateScreen("GCU Analogue Inputs", 0)
   Button "Button_16" at 550,430 size 180x50; TextOff 'Target Setpoints'; Authorization "Commissioning"
      on Press: ActivateScreen("GCU Target Setpoints", 0)
   Button "Button_17" at 550,360 size 180x50; TextOff 'Analogue Outputs'; Authorization "Commissioning"
      on Press: ActivateScreen("GCU Analogue Outputs", 0)
   Button "Button_18" at 550,500 size 180x50; TextOff 'Process Times'; Authorization "Commissioning"
      on Press: ActivateScreen("GCU Process Times", 0)
   Button "HmiScreenItemData_2" at 290,100 size 200x35; TextOn 'Back'; TextOff 'IGG Settings'
   Button "Button_7" at 300,150 size 180x50; TextOff 'Digital Inputs'; Authorization "Commissioning"
      on Click: ActivateScreen("IGG Digital Inputs", 0)
   Button "Button_8" at 300,220 size 180x50; TextOff 'Digital Outputs'; Authorization "Operating Mode"
      on Click: ActivateScreen("IGG Digital Outputs", 0)
   Button "Button_9" at 300,290 size 180x50; TextOff 'Analogue Inputs'; Authorization "Commissioning"
      on Press: ActivateScreen("IGG Analogue Inputs", 0)
   Button "Button_10" at 300,430 size 180x50; TextOff 'Target Setpoints'; Authorization "Commissioning"
      on Press: ActivateScreen("IGG Target Setpoints", 0)
   Button "Button_11" at 300,360 size 180x50; TextOff 'Analogue Outputs'; Authorization "Commissioning"
      on Press: ActivateScreen("IGG Analogue Outputs", 0)
   Button "Button_12" at 300,500 size 180x50; TextOff 'Process Times'; Authorization "Commissioning"
      on Press: ActivateScreen("IGG Process Times", 0)
   Button "HmiScreenItemData_6" at 40,100 size 200x35; TextOn 'Back'; TextOff 'BC Settings'
   Button "Button_1" at 50,150 size 180x50; TextOff 'Digital Inputs'; Authorization "Commissioning"
      on Click: ActivateScreen("BC Digital Inputs", 0)
   Button "Button_2" at 50,220 size 180x50; TextOff 'Digital Outputs'; Authorization "Operating Mode"
      on Click: ActivateScreen("BC Digital Outputs", 0)
   Button "Button_3" at 50,290 size 180x50; TextOff 'Analogue Inputs'; Authorization "Commissioning"
      on Press: ActivateScreen("BC Analogue Inputs", 0)
   Button "Button_5" at 50,430 size 180x50; TextOff 'Target Setpoints'; Authorization "Commissioning"
      on Press: ActivateScreen("BC Target Setpoints", 0)
   Button "Button_4" at 50,360 size 180x50; TextOff 'Analogue Outputs'; Authorization "Commissioning"
      on Press: ActivateScreen("BC Analogue Outputs", 0)
   Button "Button_6" at 50,570 size 180x50; TextOff 'Max Step Times'; Authorization "Commissioning"
      on Press: ActivateScreen("BC Max Step Times", 0)
   Button "HmiScreenItemData_5" at 1040,100 size 200x35; TextOn 'Back'; TextOff 'RIO Racks'
   Button "Button_25" at 1050,150 size 180x32; TextOff 'RIO 1 Digital Inputs'; Authorization "Commissioning"
      on Click: ActivateScreen("RIO 01 Digital Inputs", 0)
   Button "Button_26" at 1050,220 size 180x32; TextOff 'RIO 2 Digital Inputs'; Authorization "Operating Mode"
      on Click: ActivateScreen("RIO 02 Digital Inputs", 0)
   Button "Button_27" at 1050,290 size 180x32; TextOff 'RIO 3 Digital Inputs'; Authorization "Commissioning"
      on Click: ActivateScreen("RIO 03 Digital Inputs", 0)
   Button "Button_28" at 1050,430 size 180x32; TextOff 'RIO 5 Digital Inputs'; Authorization "Commissioning"
      on Click: ActivateScreen("RIO 05 Digital Inputs", 0)
   Button "Button_29" at 1050,360 size 180x32; TextOff 'RIO 4 Digital Inputs'; Authorization "Commissioning"
      on Click: ActivateScreen("RIO 04 Digital Inputs", 0)
   Button "Button_30" at 1050,500 size 180x32; TextOff 'RIO 6 Digital Inputs'; Authorization "Commissioning"
      on Click: ActivateScreen("RIO 06 Digital Inputs", 0)
   Button "Button_31" at 1050,570 size 180x32; TextOff 'RIO 7 Digital Inputs'; Authorization "Commissioning"
      on Click: ActivateScreen("RIO 07 Digital Inputs", 0)
   Button "Button_32" at 50,500 size 180x50; TextOff 'Process Times'; Authorization "Commissioning"
      on Press: ActivateScreen("BC Process Times", 0)
   Button "Button_33" at 300,570 size 180x50; TextOff 'Max Step Times'; Authorization "Commissioning"
      on Press: ActivateScreen("IGG Max Step Times", 0)
   Button "Button_34" at 550,570 size 180x50; TextOff 'Max Step Times'; Authorization "Commissioning"
      on Press: ActivateScreen("GCU Max Step Times", 0)
   Button "Button_19" at 1050,185 size 180x32; TextOff 'RIO 1 Analog Inputs'; Authorization "Commissioning"
      on Click: ActivateScreen("RIO 1 Analogue Settings", 0)
   Button "Button_20" at 1050,255 size 180x32; TextOff 'RIO 2 Analog Inputs'; Authorization "Operating Mode"
      on Click: ActivateScreen("RIO 2 Analogue Settings", 0)
   Button "Button_21" at 1050,325 size 180x32; TextOff 'RIO 3 Analog Inputs'; Authorization "Commissioning"
      on Click: ActivateScreen("RIO 3 Analogue Settings", 0)
   Button "Button_23" at 1050,395 size 180x32; TextOff 'RIO 4 Analog Inputs'; Authorization "Commissioning"
      on Click: ActivateScreen("RIO 4 Analogue Settings", 0)
   Button "Button_35" at 1050,465 size 180x32; TextOff 'RIO 5 Analog Inputs'; Authorization "Commissioning"
      on Click: ActivateScreen("RIO 5 Analogue Settings", 0)
   Button "Button_36" at 1050,535 size 180x32; TextOff 'RIO 6 Analog Inputs'; Authorization "Commissioning"
      on Click: ActivateScreen("RIO 6 Analogue Settings", 0)
   Button "Button_37" at 1050,604 size 180x32; TextOff 'RIO 7 Analog Inputs'; Authorization "Commissioning"
      on Click: ActivateScreen("RIO 7 Analogue Settings", 0)
   Group "Group" at 455,41 size 373x50
   Button "HmiScreenItemData_7" at 1129,1 size 150x40; TextOn 'I&A Compressor Ok'; TextOff 'Back'
      on Release: function_efd93a16()
   Button "HmiScreenItemData_8" at 469,45 size 355x40; TextOn 'Back'; TextOff 'Text'
   TextField "Screen title" at 455,41 size 373x50; Text 'Screen title'

